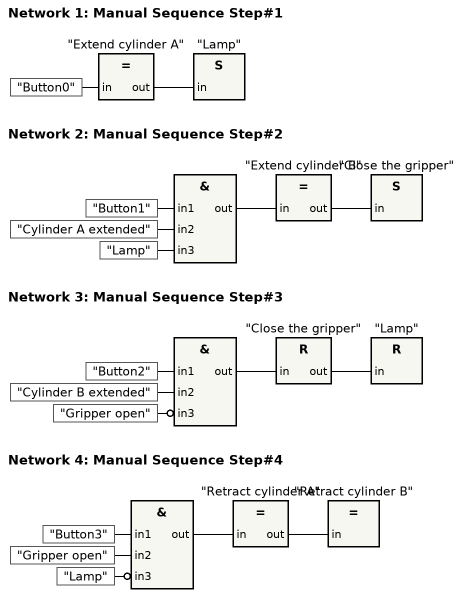
   "Extend cylinder A" := "Button0";
   IF "Button0" THEN "Lamp" := TRUE; END_IF;
END_REGION

REGION Network 2: Manual Sequence Step#2
   // Pressing button I1.1 extends cylinder B and closes the gripper
   "Extend cylinder B" := "Button1" AND "Cylinder A extended" AND "Lamp";
   IF "Extend cylinder B" THEN "Close the gripper" := TRUE; END_IF;
END_REGION

REGION Network 3: Manual Sequence Step#3
   // Pressing button I1.2 opens the gripper and turns the lamp OFF
   IF "Button2" AND "Cylinder B extended" AND NOT "Gripper open" THEN
       "Close the gripper" := FALSE;
       "Lamp" := FALSE;
   END_IF;
END_REGION

REGION Network 4: Manual Sequence Step#4
   // Pressing button I1.3 retracts the cylinders
   "Retract cylinder A" := "Button3" AND "Gripper open" AND NOT "Lamp";
   "Retract cylinder B" := "Retract cylinder A";
END_REGION
END_FUNCTION

FUNCTION "FC020_Three_Production_Lines" : Void   // FC25, LAD
{ S7_Optimized_Access := 'TRUE' }
VERSION : 0.1
   VAR_TEMP   // added for the SCL form of the ladder/FBD networks
      _w1 : Bool;
   END_VAR
BEGIN

REGION Network 1: Counters Reset
   // Button OFF resets Line 1, Line 2, Line 3 quantity counters and the Total Profit value
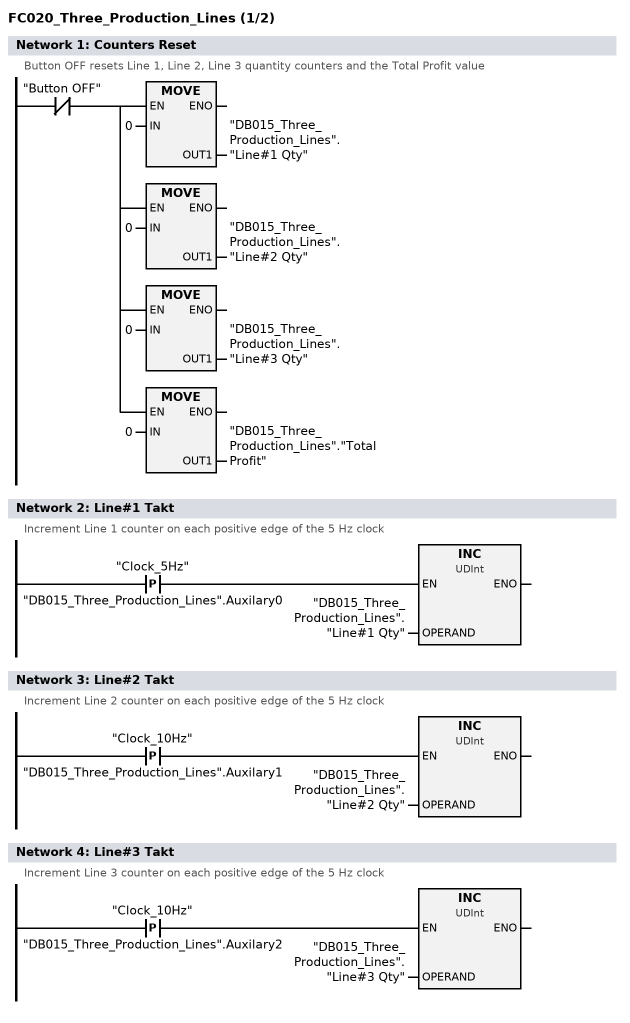
   RUNG wire#powerrail
      I_Contact( "Button OFF" )
      wire#w1
      Move(in := 0, out1 => "DB015_Three_Production_Lines"."Line#1 Qty")
   END_RUNG
   RUNG wire#w1
      Move(in := 0, out1 => "DB015_Three_Production_Lines"."Line#2 Qty")
   END_RUNG
   RUNG wire#w1
      Move(in := 0, out1 => "DB015_Three_Production_Lines"."Line#3 Qty")
   END_RUNG
   RUNG wire#w1
      Move(in := 0, out1 => "DB015_Three_Production_Lines"."Total Profit")
   END_RUNG
   // the same network as SCL:
   IF NOT "Button OFF" THEN
       "DB015_Three_Production_Lines"."Line#1 Qty" := 0;
       "DB015_Three_Production_Lines"."Line#2 Qty" := 0;
       "DB015_Three_Production_Lines"."Line#3 Qty" := 0;
       "DB015_Three_Production_Lines"."Total Profit" := 0;
   END_IF;
END_REGION

REGION Network 2: Line#1 Takt
   // Increment Line 1 counter on each positive edge of the 5 Hz clock
   RUNG wire#powerrail
      P_Contact(operand := "Clock_5Hz", bit := "DB015_Three_Production_Lines".Auxilary0)
      { S7_Templates := "DestType := UDInt" } Inc( "DB015_Three_Production_Lines"."Line#1 Qty" )
   END_RUNG
   // the same network as SCL:
   #_w1 := "Clock_5Hz" AND NOT "DB015_Three_Production_Lines".Auxilary0;   // rising edge of "Clock_5Hz"
   "DB015_Three_Production_Lines".Auxilary0 := "Clock_5Hz";
   IF #_w1 THEN
       "DB015_Three_Production_Lines"."Line#1 Qty" := "DB015_Three_Production_Lines"."Line#1 Qty" + 1;
   END_IF;
END_REGION

REGION Network 3: Line#2 Takt
   // Increment Line 2 counter on each positive edge of the 5 Hz clock
   RUNG wire#powerrail
      P_Contact(operand := "Clock_10Hz", bit := "DB015_Three_Production_Lines".Auxilary1)
      { S7_Templates := "DestType := UDInt" } Inc( "DB015_Three_Production_Lines"."Line#2 Qty" )
   END_RUNG
   // the same network as SCL:
   #_w1 := "Clock_10Hz" AND NOT "DB015_Three_Production_Lines".Auxilary1;   // rising edge of "Clock_10Hz"
   "DB015_Three_Production_Lines".Auxilary1 := "Clock_10Hz";
   IF #_w1 THEN
       "DB015_Three_Production_Lines"."Line#2 Qty" := "DB015_Three_Production_Lines"."Line#2 Qty" + 1;
   END_IF;
END_REGION

REGION Network 4: Line#3 Takt
   // Increment Line 3 counter on each positive edge of the 5 Hz clock
   RUNG wire#powerrail
      P_Contact(operand := "Clock_10Hz", bit := "DB015_Three_Production_Lines".Auxilary2)
      { S7_Templates := "DestType := UDInt" } Inc( "DB015_Three_Production_Lines"."Line#3 Qty" )
   END_RUNG
   // the same network as SCL:
   #_w1 := "Clock_10Hz" AND NOT "DB015_Three_Production_Lines".Auxilary2;   // rising edge of "Clock_10Hz"
   "DB015_Three_Production_Lines".Auxilary2 := "Clock_10Hz";
   IF #_w1 THEN
       "DB015_Three_Production_Lines"."Line#3 Qty" := "DB015_Three_Production_Lines"."Line#3 Qty" + 1;
   END_IF;
END_REGION

REGION Network 5: Current Profit Calculation
   // Calculate the current profit as a weighted sum: Profit=L1_Qty*Price1+L2_Qty*Price2+L3_Qty*Price3
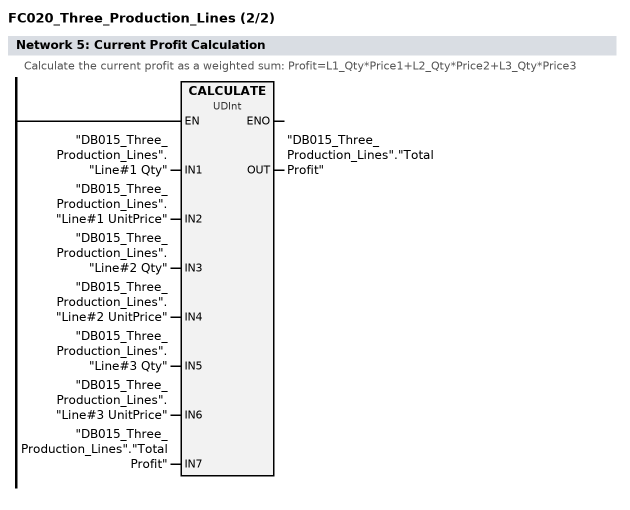
   RUNG wire#powerrail
      { S7_Templates := "SrcType := UDInt"; S7_Expression := "IN7 + (IN1 * IN2 + IN3 * IN4 + IN5 * IN6)" } Calculate(in1 := "DB015_Three_Production_Lines"."Line#1 Qty", in2 := "DB015_Three_Production_Lines"."Line#1 UnitPrice", in3 := "DB015_Three_Production_Lines"."Line#2 Qty", in4 := "DB015_Three_Production_Lines"."Line#2 UnitPrice", in5 := "DB015_Three_Production_Lines"."Line#3 Qty", in6 := "DB015_Three_Production_Lines"."Line#3 UnitPrice", in7 := "DB015_Three_Production_Lines"."Total Profit", out => "DB015_Three_Production_Lines"."Total Profit")
   END_RUNG
   // the same network as SCL:
   "DB015_Three_Production_Lines"."Total Profit" := "DB015_Three_Production_Lines"."Total Profit" + ("DB015_Three_Production_Lines"."Line#1 Qty" * "DB015_Three_Production_Lines"."Line#1 UnitPrice" + "DB015_Three_Production_Lines"."Line#2 Qty" * "DB015_Three_Production_Lines"."Line#2 UnitPrice" + "DB015_Three_Production_Lines"."Line#3 Qty" * "DB015_Three_Production_Lines"."Line#3 UnitPrice");
END_REGION
END_FUNCTION

FUNCTION "FC021_Packaging_Control" : Void   // FC26, LAD
{ S7_Optimized_Access := 'TRUE' }
VERSION : 0.1
BEGIN

REGION Network 1: Bottle, Row, and Box Counting Logic
   // Every 1s pulse increments the bottle counter. 
   // Reaching 4 bottles triggers Next Row and resets the bottle counter. 
   // Next Row increments the row counter. 
   // Reaching 6 rows triggers Next Box, resetting the row counter and incrementing the box counter (INC).
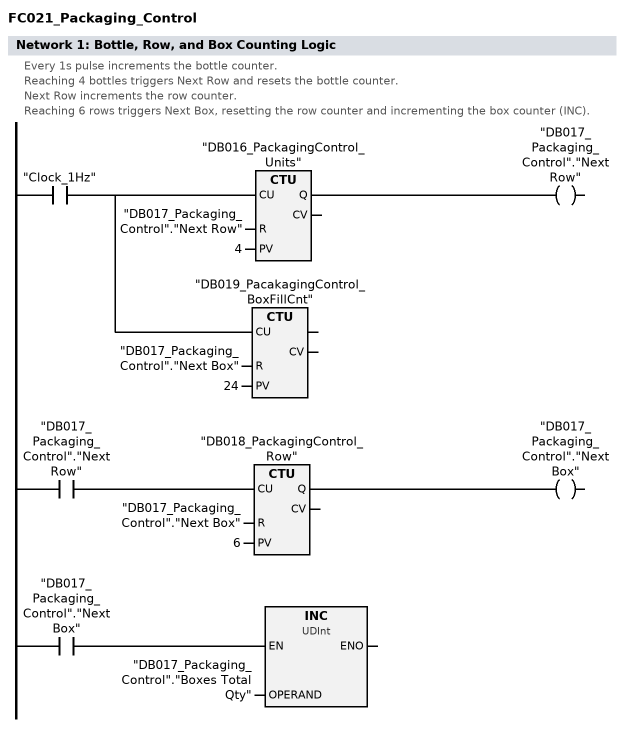
   "DB016_PackagingControl_Units".CTU(CU := "Clock_1Hz", R := "DB017_Packaging_Control"."Next Row", PV := 4);
   "DB017_Packaging_Control"."Next Row" := "DB016_PackagingControl_Units".Q;
   "DB019_PacakagingControl_BoxFillCnt".CTU(CU := "Clock_1Hz",
                           R := "DB017_Packaging_Control"."Next Box",
                           PV := 24);
   "DB018_PackagingControl_Row".CTU(CU := "DB017_Packaging_Control"."Next Row",
                           R := "DB017_Packaging_Control"."Next Box",
                           PV := 6);
   "DB017_Packaging_Control"."Next Box" := "DB018_PackagingControl_Row".Q;
   IF "DB017_Packaging_Control"."Next Box" THEN
       "DB017_Packaging_Control"."Boxes Total Qty" := "DB017_Packaging_Control"."Boxes Total Qty" + 1;
   END_IF;
END_REGION
END_FUNCTION

ORGANIZATION_BLOCK "Main"   // OB1, LAD, ProgramCycle
TITLE = "Main Program Sweep (Cycle)"
{ S7_Optimized_Access := 'TRUE' }
VERSION : 0.1
   VAR_INPUT
      Initial_Call : Bool;   // Initial call of this OB
      Remanence : Bool;   // =True, if remanent data are available
   END_VAR
BEGIN
END_ORGANIZATION_BLOCK

(* ===== HMI "HMI_RT_1" =====
system functions are stored by id; their names below are inferred from use
connection "HMI_Connection_1": ETHERNET, SMART_S7_1200_OMS

HMI tags "HMI Tags"
   "DB002_Auto_Cycle_HMI_Start" : Bool = PLC DB002_Auto_Cycle.HMI_Start, 1 s
   "DB002_Auto_Cycle_HMI_Stop" : Bool = PLC DB002_Auto_Cycle.HMI_Stop AT %DB1.DBX0.0, 1 s
   "Clock_1Hz" : Bool = PLC Clock_1Hz AT %M0.5, 1 s
   "Cylinder A extended" : Bool = PLC "Cylinder A extended" AT %I0.6, 1 s
   "Cylinder B extended" : Bool = PLC "Cylinder B extended" AT %I0.4, 1 s
   "Gripper open" : Bool = PLC "Gripper open" AT %I0.5, 1 s
   "DB004_Labeler_Control_Labels_Counter" : Int = PLC DB004_Labeler_Control.Labels_Counter, 1 s
   "DB004_Labeler_Control_Number_of_Labels_Remaining" : Int = PLC DB004_Labeler_Control.Number_of_Labels_Remaining, 1 s
   "DB004_Labeler_Control_Label_Rolls_Counter" : Int = PLC DB004_Labeler_Control.Label_Rolls_Counter, 1 s

Template "Template_1" 800x480
   Button "Exit" at 714,429 size 71x50; TextOff 'Exit'; PictureOff "ExitRuntime_KTP700_Basic_PN_TR"; PictureOn "ExitRuntime_KTP700_Basic_PN_TR"
      on Release: StopRuntime(0)
   Button "Language" at 614,429 size 71x50; TextOff 'Language'; PictureOff "ToggleLanguage_KTP700_Basic_PN_TR"; PictureOn "ToggleLanguage_KTP700_Basic_PN_TR"
      on Release: function_fb9197e8(-1)
   Button "Template_Button" at 514,429 size 71x50; TextOff 'Text'
   Button "Template_Button_1" at 414,429 size 71x50; TextOff 'Text'
   Button "Template_Button_2" at 314,429 size 71x50; TextOff 'Text'
   Button "Log on" at 214,429 size 71x50; TextOff 'Log on'; PictureOff "Login_KTP700_Basic_PN_TR"; PictureOn "Login_KTP700_Basic_PN_TR"
      on Release: function_a2a04561()
   Button "Alarms" at 114,429 size 71x50; TextOff 'Alarms'; PictureOff "AlarmDisplay_KTP700_Basic_PN_TR"; PictureOn "AlarmDisplay_KTP700_Basic_PN_TR"
      on Release: function_ef3f5d25("Alarm window_Unacknowledged", -1)
   Button "Start screen" at 14,429 size 71x50; TextOff 'Start screen'; PictureOff "NavigateHome_KTP700_Basic_PN_TR"; PictureOn "NavigateHome_KTP700_Basic_PN_TR"
      on Release: ActivateScreen("Home", 0)
   SymbolicIOField "Symbolic_IO_Field_Screen" at 93,9 size 600x33; TextOff '0'; TextOn '1'; TextList "TextList_ScreenNames"
      ProcessValue <- "Tag_ScreenNumber"
      on Change: ActivateScreenByNumber("Tag_ScreenNumber", 0)
   DateTimeField "HmiScreenItemData" at 695,25 size 105x25
   DateTimeField "HmiScreenItemData_1" at 695,0 size 105x25
   GraphicView "Logo" at 0,0 size 91x51; Picture "Logo of HMI_1"

screen "Home" 800x480, template "Template_1"
   on GenerateScreen: SetTag("Tag_ScreenNumber", 1)
   Circle "Circle_1" at 708,76 size 67x67
      Appearance <- "Clock_1Hz"
   TextField "Text field_1" at 86,65 size 171x23; Text 'Cylinder A Extended'
   TextField "Text field_2" at 87,102 size 170x23; Text 'Cylinder B Extended'
   Rectangle "Rectangle_1" at 272,60 size 32x28
      Appearance <- "Cylinder A extended"
   Rectangle "Rectangle_2" at 272,97 size 32x28
      Appearance <- "Cylinder B extended"
   Rectangle "Rectangle_3" at 272,135 size 32x28
      Appearance <- "Gripper open"
   TextField "Text field_3" at 87,140 size 133x23; Text 'Gripper Opened'
   Button "Button_1" at 223,359 size 155x52; TextOff 'CYCLE START'
      on Press: function_b14e0dd5("DB002_Auto_Cycle_HMI_Start", 0)
   Button "Button_2" at 424,359 size 155x52; TextOff 'CYCLE STOP'
      on Press: function_b14e0dd5("DB002_Auto_Cycle_HMI_Stop", 0)
   IOField "I/O field_1" at 358,194 size 96x32; FormatPattern 999
      ProcessValue <- "DB004_Labeler_Control_Labels_Counter"
   TextField "Text field_4" at 116,196 size 144x23; Text 'Bottles Produced'
   IOField "I/O field_2" at 358,239 size 96x32; FormatPattern 999
      ProcessValue <- "DB004_Labeler_Control_Number_of_Labels_Remaining"
   TextField "Text field_5" at 116,239 size 149x23; Text 'Labels Remaining'
   IOField "I/O field_3" at 358,286 size 96x32; FormatPattern 999
      ProcessValue <- "DB004_Labeler_Control_Label_Rolls_Counter"
   TextField "Text field_6" at 116,286 size 180x23; Text 'Number of Rolls Used'
*)